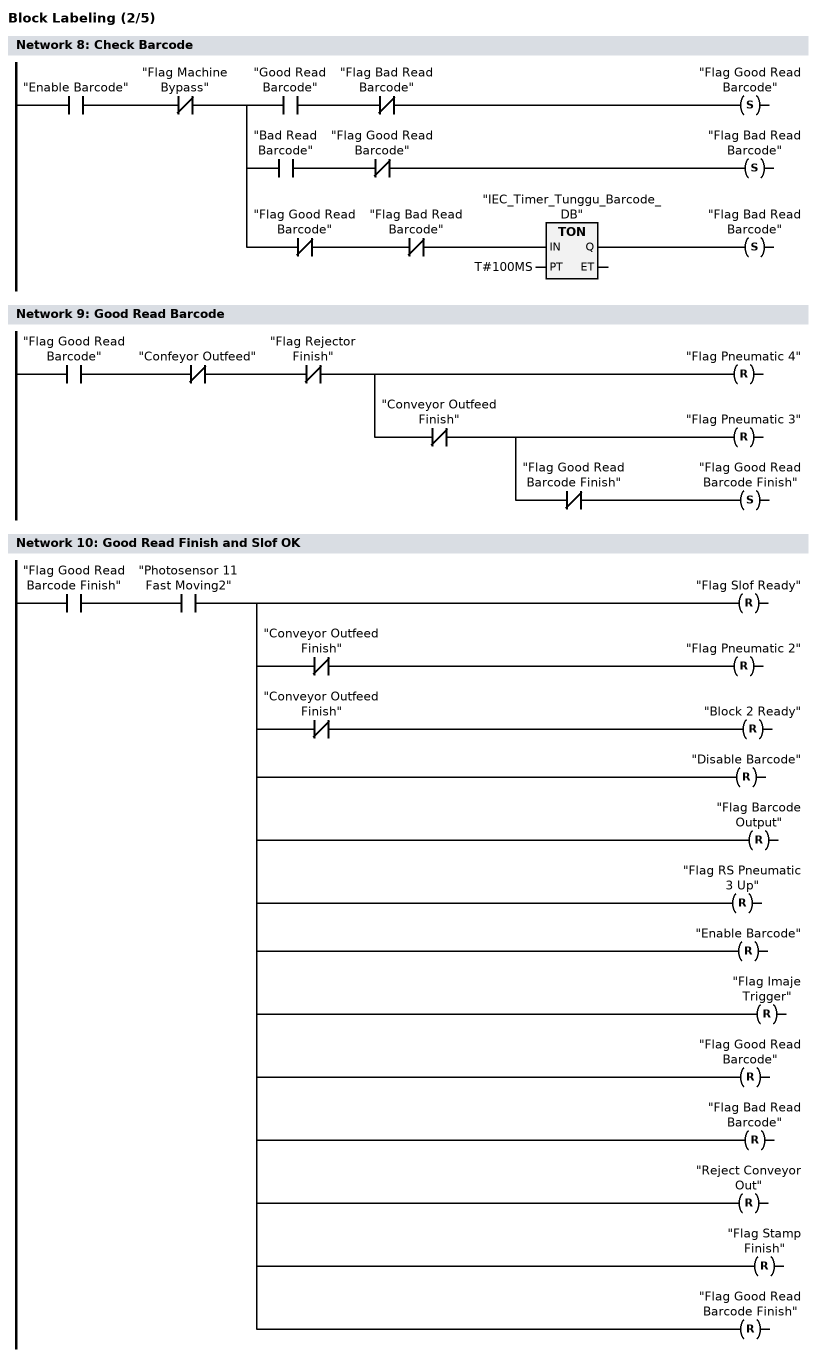
   #_w1 := "Enable Barcode" AND NOT "Flag Machine Bypass";
   IF #_w1 AND "Good Read Barcode" AND NOT "Flag Bad Read Barcode" THEN
       "Flag Good Read Barcode" := TRUE;
   END_IF;
   IF #_w1 AND "Bad Read Barcode" AND NOT "Flag Good Read Barcode" THEN
       "Flag Bad Read Barcode" := TRUE;
   END_IF;
   "IEC_Timer_Tunggu_Barcode_DB".TON(IN := #_w1 AND NOT "Flag Good Read Barcode" AND NOT "Flag Bad Read Barcode",
                           PT := T#100MS);
   IF "IEC_Timer_Tunggu_Barcode_DB".Q THEN "Flag Bad Read Barcode" := TRUE; END_IF;
END_REGION

REGION Network 9: Good Read Barcode
   RUNG wire#powerrail
      Contact( "Flag Good Read Barcode" )
      I_Contact( "Confeyor Outfeed" )
      I_Contact( "Flag Rejector Finish" )
      wire#w1
      R_Coil( "Flag Pneumatic 4" )
   END_RUNG
   RUNG wire#w1
      I_Contact( "Conveyor Outfeed Finish" )
      wire#w2
      R_Coil( "Flag Pneumatic 3" )
   END_RUNG
   RUNG wire#w2
      I_Contact( "Flag Good Read Barcode Finish" )
      S_Coil( "Flag Good Read Barcode Finish" )
   END_RUNG
   // the same network as SCL:
   #_w1 := "Flag Good Read Barcode" AND NOT "Confeyor Outfeed" AND NOT "Flag Rejector Finish";
   IF #_w1 THEN "Flag Pneumatic 4" := FALSE; END_IF;
   #_w2 := #_w1 AND NOT "Conveyor Outfeed Finish";
   IF #_w2 THEN "Flag Pneumatic 3" := FALSE; END_IF;
   IF #_w2 AND NOT "Flag Good Read Barcode Finish" THEN "Flag Good Read Barcode Finish" := TRUE; END_IF;
END_REGION

REGION Network 10: Good Read Finish and Slof OK
   RUNG wire#powerrail
      Contact( "Flag Good Read Barcode Finish" )
      Contact( "Photosensor 11 Fast Moving2" )
      wire#w1
      R_Coil( "Flag Slof Ready" )
   END_RUNG
   RUNG wire#w1
      I_Contact( "Conveyor Outfeed Finish" )
      R_Coil( "Flag Pneumatic 2" )
   END_RUNG
   RUNG wire#w1
      I_Contact( "Conveyor Outfeed Finish" )
      R_Coil( "Block 2 Ready" )
   END_RUNG
   RUNG wire#w1
      R_Coil( "Disable Barcode" )
   END_RUNG
   RUNG wire#w1
      R_Coil( "Flag Barcode Output" )
   END_RUNG
   RUNG wire#w1
      R_Coil( "Flag RS Pneumatic 3 Up" )
   END_RUNG
   RUNG wire#w1
      R_Coil( "Enable Barcode" )
   END_RUNG
   RUNG wire#w1
      R_Coil( "Flag Imaje Trigger" )
   END_RUNG
   RUNG wire#w1
      R_Coil( "Flag Good Read Barcode" )
   END_RUNG
   RUNG wire#w1
      R_Coil( "Flag Bad Read Barcode" )
   END_RUNG
   RUNG wire#w1
      R_Coil( "Reject Conveyor Out" )
   END_RUNG
   RUNG wire#w1
      R_Coil( "Flag Stamp Finish" )
   END_RUNG
   RUNG wire#w1
      R_Coil( "Flag Good Read Barcode Finish" )
   END_RUNG
   // the same network as SCL:
   #_w1 := "Flag Good Read Barcode Finish" AND "Photosensor 11 Fast Moving2";
   IF #_w1 THEN "Flag Slof Ready" := FALSE; END_IF;
   IF #_w1 AND NOT "Conveyor Outfeed Finish" THEN
       "Flag Pneumatic 2" := FALSE;
       "Block 2 Ready" := FALSE;
   END_IF;
   IF #_w1 THEN
       "Disable Barcode" := FALSE;
       "Flag Barcode Output" := FALSE;
       "Flag RS Pneumatic 3 Up" := FALSE;
       "Enable Barcode" := FALSE;
       "Flag Imaje Trigger" := FALSE;
       "Flag Good Read Barcode" := FALSE;
       "Flag Bad Read Barcode" := FALSE;
       "Reject Conveyor Out" := FALSE;
       "Flag Stamp Finish" := FALSE;
       "Flag Good Read Barcode Finish" := FALSE;
   END_IF;
END_REGION

REGION Network 11: Set Section Reject
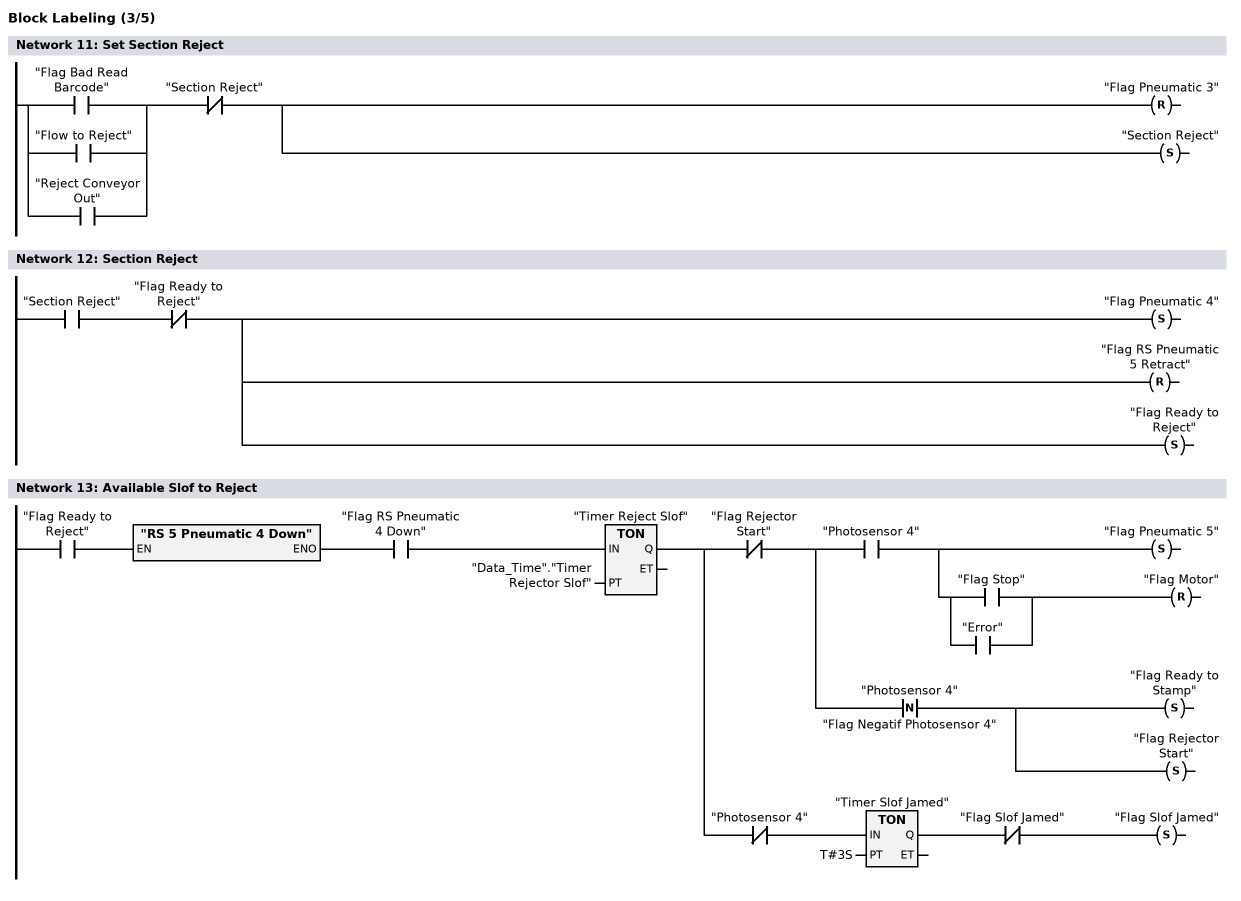
   RUNG wire#powerrail
      Contact( "Flag Bad Read Barcode" )
      wire#w1
      I_Contact( "Section Reject" )
      wire#w2
      R_Coil( "Flag Pneumatic 3" )
   END_RUNG
   RUNG wire#powerrail
      Contact( "Flow to Reject" )
   END_RUNG wire#w1
   RUNG wire#powerrail
      Contact( "Reject Conveyor Out" )
   END_RUNG wire#w1
   RUNG wire#w2
      S_Coil( "Section Reject" )
   END_RUNG
   // the same network as SCL:
   IF ("Flag Bad Read Barcode" OR "Flow to Reject" OR "Reject Conveyor Out") AND NOT "Section Reject" THEN
       "Flag Pneumatic 3" := FALSE;
       "Section Reject" := TRUE;
   END_IF;
END_REGION

REGION Network 12: Section Reject
   RUNG wire#powerrail
      Contact( "Section Reject" )
      I_Contact( "Flag Ready to Reject" )
      wire#w1
      S_Coil( "Flag Pneumatic 4" )
   END_RUNG
   RUNG wire#w1
      R_Coil( "Flag RS Pneumatic 5 Retract" )
   END_RUNG
   RUNG wire#w1
      S_Coil( "Flag Ready to Reject" )
   END_RUNG
   // the same network as SCL:
   IF "Section Reject" AND NOT "Flag Ready to Reject" THEN
       "Flag Pneumatic 4" := TRUE;
       "Flag RS Pneumatic 5 Retract" := FALSE;
       "Flag Ready to Reject" := TRUE;
   END_IF;
END_REGION

REGION Network 13: Available Slof to Reject
   "RS 5 Pneumatic 4 Down"(EN := "Flag Ready to Reject", ENO => #_w1);
   "Timer Reject Slof".TON(IN := #_w1 AND "Flag RS Pneumatic 4 Down", PT := "Data_Time"."Timer Rejector Slof");
   #_w2 := "Timer Reject Slof".Q AND NOT "Flag Rejector Start";
   #_w3 := #_w2 AND "Photosensor 4";
   IF #_w3 THEN "Flag Pneumatic 5" := TRUE; END_IF;
   IF #_w3 AND ("Flag Stop" OR "Error") THEN "Flag Motor" := FALSE; END_IF;
   #_w4 := #_w2 AND NOT "Photosensor 4" AND "Flag Negatif Photosensor 4";   // falling edge of "Photosensor 4"
   "Flag Negatif Photosensor 4" := "Photosensor 4";
   IF #_w4 THEN
       "Flag Ready to Stamp" := TRUE;
       "Flag Rejector Start" := TRUE;
   END_IF;
   "Timer Slof Jamed".TON(IN := "Timer Reject Slof".Q AND NOT "Photosensor 4", PT := T#3S);
   IF "Timer Slof Jamed".Q AND NOT "Flag Slof Jamed" THEN "Flag Slof Jamed" := TRUE; END_IF;
END_REGION

REGION Network 14: Ready to Stamp again
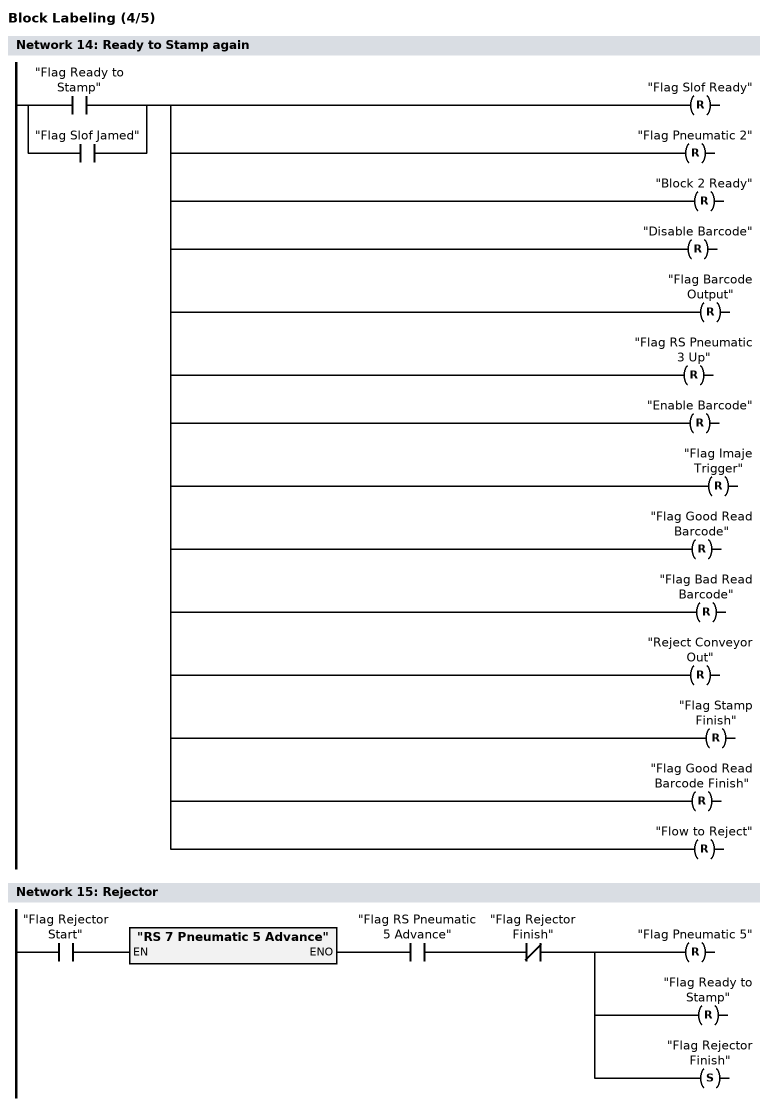
   RUNG wire#powerrail
      Contact( "Flag Ready to Stamp" )
      wire#w1
      R_Coil( "Flag Slof Ready" )
   END_RUNG
   RUNG wire#powerrail
      Contact( "Flag Slof Jamed" )
   END_RUNG wire#w1
   RUNG wire#w1
      R_Coil( "Flag Pneumatic 2" )
   END_RUNG
   RUNG wire#w1
      R_Coil( "Block 2 Ready" )
   END_RUNG
   RUNG wire#w1
      R_Coil( "Disable Barcode" )
   END_RUNG
   RUNG wire#w1
      R_Coil( "Flag Barcode Output" )
   END_RUNG
   RUNG wire#w1
      R_Coil( "Flag RS Pneumatic 3 Up" )
   END_RUNG
   RUNG wire#w1
      R_Coil( "Enable Barcode" )
   END_RUNG
   RUNG wire#w1
      R_Coil( "Flag Imaje Trigger" )
   END_RUNG
   RUNG wire#w1
      R_Coil( "Flag Good Read Barcode" )
   END_RUNG
   RUNG wire#w1
      R_Coil( "Flag Bad Read Barcode" )
   END_RUNG
   RUNG wire#w1
      R_Coil( "Reject Conveyor Out" )
   END_RUNG
   RUNG wire#w1
      R_Coil( "Flag Stamp Finish" )
   END_RUNG
   RUNG wire#w1
      R_Coil( "Flag Good Read Barcode Finish" )
   END_RUNG
   RUNG wire#w1
      R_Coil( "Flow to Reject" )
   END_RUNG
   // the same network as SCL:
   IF "Flag Ready to Stamp" OR "Flag Slof Jamed" THEN
       "Flag Slof Ready" := FALSE;
       "Flag Pneumatic 2" := FALSE;
       "Block 2 Ready" := FALSE;
       "Disable Barcode" := FALSE;
       "Flag Barcode Output" := FALSE;
       "Flag RS Pneumatic 3 Up" := FALSE;
       "Enable Barcode" := FALSE;
       "Flag Imaje Trigger" := FALSE;
       "Flag Good Read Barcode" := FALSE;
       "Flag Bad Read Barcode" := FALSE;
       "Reject Conveyor Out" := FALSE;
       "Flag Stamp Finish" := FALSE;
       "Flag Good Read Barcode Finish" := FALSE;
       "Flow to Reject" := FALSE;
   END_IF;
END_REGION

REGION Network 15: Rejector
   RUNG wire#powerrail
      Contact( "Flag Rejector Start" )
      "RS 7 Pneumatic 5 Advance"()
      Contact( "Flag RS Pneumatic 5 Advance" )
      I_Contact( "Flag Rejector Finish" )
      wire#w1
      R_Coil( "Flag Pneumatic 5" )
   END_RUNG
   RUNG wire#w1
      R_Coil( "Flag Ready to Stamp" )
   END_RUNG
   RUNG wire#w1
      S_Coil( "Flag Rejector Finish" )
   END_RUNG
   // the same network as SCL:
   "RS 7 Pneumatic 5 Advance"(EN := "Flag Rejector Start", ENO => #_w1);
   IF #_w1 AND "Flag RS Pneumatic 5 Advance" AND NOT "Flag Rejector Finish" THEN
       "Flag Pneumatic 5" := FALSE;
       "Flag Ready to Stamp" := FALSE;
       "Flag Rejector Finish" := TRUE;
   END_IF;
END_REGION

REGION Network 16: Rejector Finish
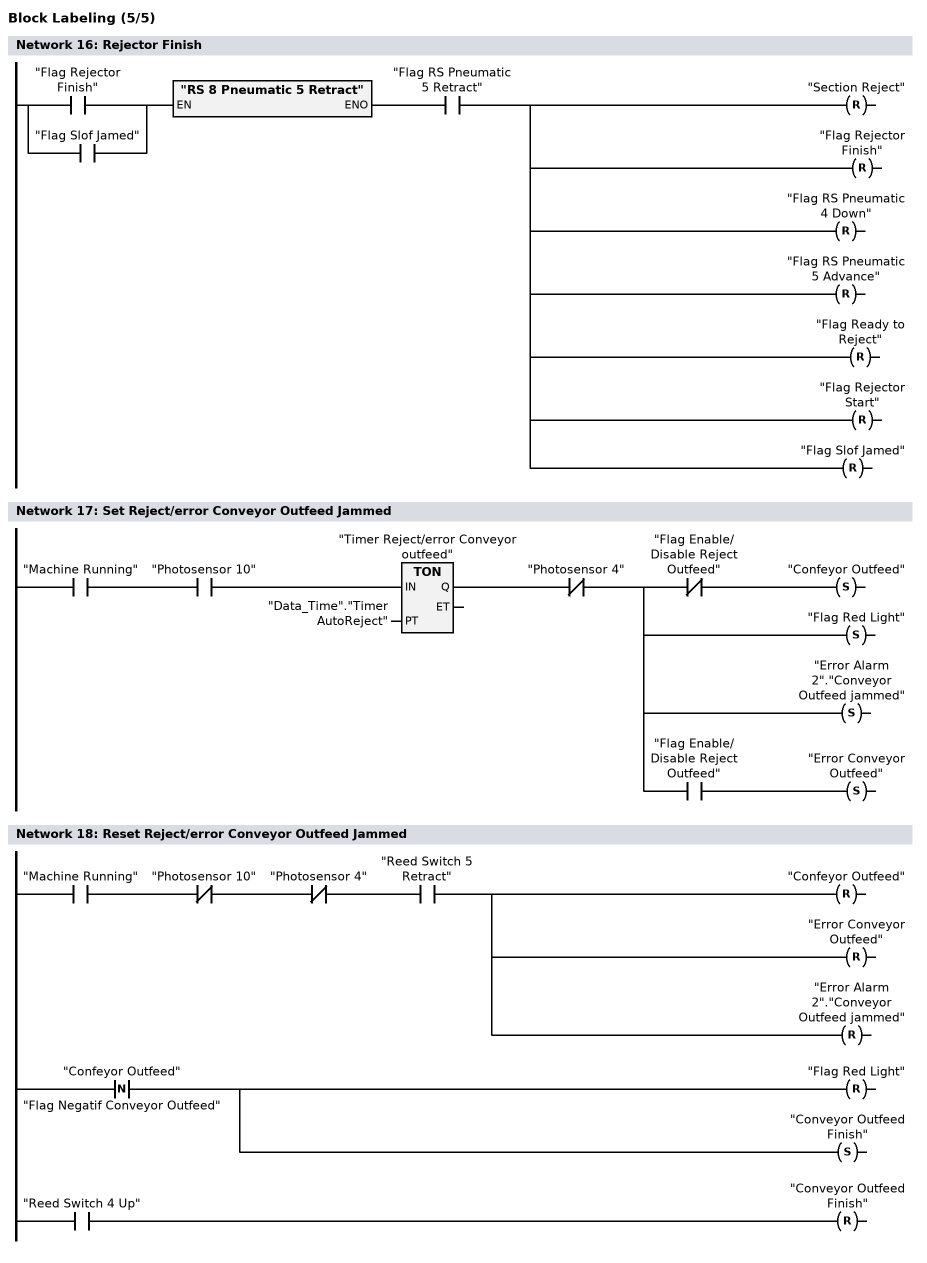
   RUNG wire#powerrail
      Contact( "Flag Rejector Finish" )
      wire#w1
      "RS 8 Pneumatic 5 Retract"()
      Contact( "Flag RS Pneumatic 5 Retract" )
      wire#w2
      R_Coil( "Section Reject" )
   END_RUNG
   RUNG wire#powerrail
      Contact( "Flag Slof Jamed" )
   END_RUNG wire#w1
   RUNG wire#w2
      R_Coil( "Flag Rejector Finish" )
   END_RUNG
   RUNG wire#w2
      R_Coil( "Flag RS Pneumatic 4 Down" )
   END_RUNG
   RUNG wire#w2
      R_Coil( "Flag RS Pneumatic 5 Advance" )
   END_RUNG
   RUNG wire#w2
      R_Coil( "Flag Ready to Reject" )
   END_RUNG
   RUNG wire#w2
      R_Coil( "Flag Rejector Start" )
   END_RUNG
   RUNG wire#w2
      R_Coil( "Flag Slof Jamed" )
   END_RUNG
   // the same network as SCL:
   "RS 8 Pneumatic 5 Retract"(EN := "Flag Rejector Finish" OR "Flag Slof Jamed", ENO => #_w1);
   IF #_w1 AND "Flag RS Pneumatic 5 Retract" THEN
       "Section Reject" := FALSE;
       "Flag Rejector Finish" := FALSE;
       "Flag RS Pneumatic 4 Down" := FALSE;
       "Flag RS Pneumatic 5 Advance" := FALSE;
       "Flag Ready to Reject" := FALSE;
       "Flag Rejector Start" := FALSE;
       "Flag Slof Jamed" := FALSE;
   END_IF;
END_REGION

REGION Network 17: Set Reject/error Conveyor Outfeed Jammed
   "Timer Reject/error Conveyor outfeed".TON(IN := "Machine Running" AND "Photosensor 10",
                           PT := "Data_Time"."Timer AutoReject");
   #_w1 := "Timer Reject/error Conveyor outfeed".Q AND NOT "Photosensor 4";
   IF #_w1 AND NOT "Flag Enable/Disable Reject Outfeed" THEN "Confeyor Outfeed" := TRUE; END_IF;
   IF #_w1 THEN
       "Flag Red Light" := TRUE;
       "Error Alarm 2"."Conveyor Outfeed jammed" := TRUE;
   END_IF;
   IF #_w1 AND "Flag Enable/Disable Reject Outfeed" THEN "Error Conveyor Outfeed" := TRUE; END_IF;
END_REGION

REGION Network 18: Reset Reject/error Conveyor Outfeed Jammed
   RUNG wire#powerrail
      Contact( "Machine Running" )
      I_Contact( "Photosensor 10" )
      I_Contact( "Photosensor 4" )
      Contact( "Reed Switch 5 Retract" )
      wire#w1
      R_Coil( "Confeyor Outfeed" )
   END_RUNG
   RUNG wire#w1
      R_Coil( "Error Conveyor Outfeed" )
   END_RUNG
   RUNG wire#w1
      R_Coil( "Error Alarm 2"."Conveyor Outfeed jammed" )
   END_RUNG
   RUNG wire#powerrail
      N_Contact(operand := "Confeyor Outfeed", bit := "Flag Negatif Conveyor Outfeed")
      wire#w2
      R_Coil( "Flag Red Light" )
   END_RUNG
   RUNG wire#w2
      S_Coil( "Conveyor Outfeed Finish" )
   END_RUNG
   RUNG wire#powerrail
      Contact( "Reed Switch 4 Up" )
      R_Coil( "Conveyor Outfeed Finish" )
   END_RUNG
   // the same network as SCL:
   IF "Machine Running" AND NOT "Photosensor 10" AND NOT "Photosensor 4" AND "Reed Switch 5 Retract" THEN
       "Confeyor Outfeed" := FALSE;
       "Error Conveyor Outfeed" := FALSE;
       "Error Alarm 2"."Conveyor Outfeed jammed" := FALSE;
   END_IF;
   #_w1 := NOT "Confeyor Outfeed" AND "Flag Negatif Conveyor Outfeed";   // falling edge of "Confeyor Outfeed"
   "Flag Negatif Conveyor Outfeed" := "Confeyor Outfeed";
   IF #_w1 THEN
       "Flag Red Light" := FALSE;
       "Conveyor Outfeed Finish" := TRUE;
   END_IF;
   IF "Reed Switch 4 Up" THEN "Conveyor Outfeed Finish" := FALSE; END_IF;
END_REGION
END_FUNCTION_BLOCK

FUNCTION_BLOCK "Block Focke"   // FB6, LAD
{ S7_Optimized_Access := 'TRUE' }
VERSION : 0.1
   VAR_TEMP   // added for the SCL form of the ladder/FBD networks
      _w1 : Bool;
   END_VAR
BEGIN

REGION Network 1: Enable/Disable Error Chute Before Heating Roll
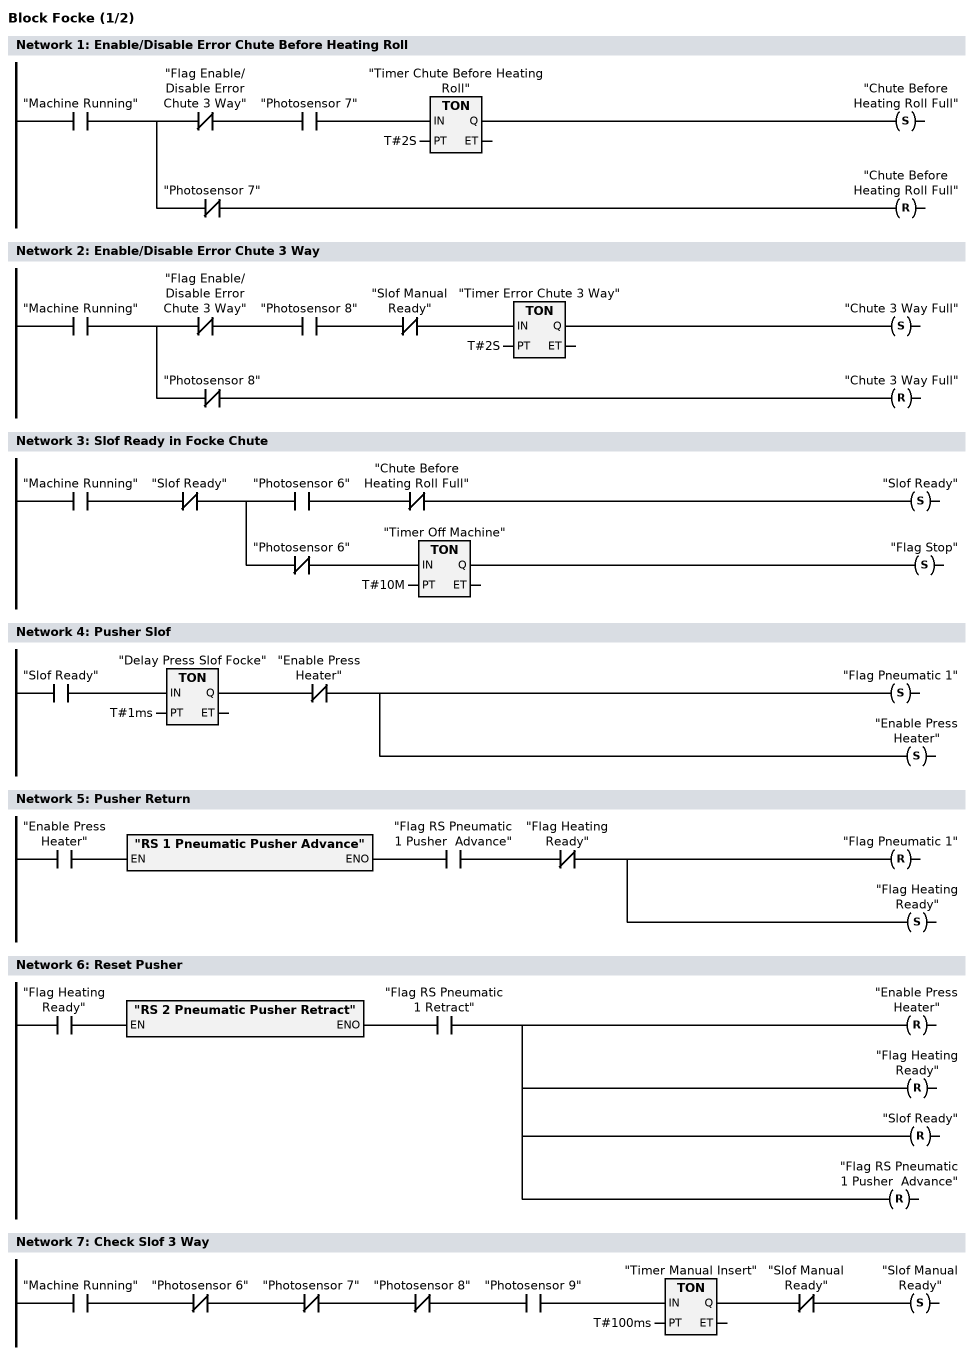
   "Timer Chute Before Heating Roll".TON(IN := "Machine Running" AND NOT "Flag Enable/Disable Error Chute 3 Way" AND "Photosensor 7",
                           PT := T#2S);
   IF "Timer Chute Before Heating Roll".Q THEN "Chute Before Heating Roll Full" := TRUE; END_IF;
   IF "Machine Running" AND NOT "Photosensor 7" THEN "Chute Before Heating Roll Full" := FALSE; END_IF;
END_REGION

REGION Network 2: Enable/Disable Error Chute 3 Way
   "Timer Error Chute 3 Way".TON(IN := "Machine Running" AND NOT "Flag Enable/Disable Error Chute 3 Way" AND "Photosensor 8" AND NOT "Slof Manual Ready",
                           PT := T#2S);
   IF "Timer Error Chute 3 Way".Q THEN "Chute 3 Way Full" := TRUE; END_IF;
   IF "Machine Running" AND NOT "Photosensor 8" THEN "Chute 3 Way Full" := FALSE; END_IF;
END_REGION

REGION Network 3: Slof Ready in Focke Chute
   #_w1 := "Machine Running" AND NOT "Slof Ready";
   IF #_w1 AND "Photosensor 6" AND NOT "Chute Before Heating Roll Full" THEN "Slof Ready" := TRUE; END_IF;
   "Timer Off Machine".TON(IN := #_w1 AND NOT "Photosensor 6", PT := T#10M);
   IF "Timer Off Machine".Q THEN "Flag Stop" := TRUE; END_IF;
END_REGION

REGION Network 4: Pusher Slof
   "Delay Press Slof Focke".TON(IN := "Slof Ready", PT := T#1ms);
   IF "Delay Press Slof Focke".Q AND NOT "Enable Press Heater" THEN
       "Flag Pneumatic 1" := TRUE;
       "Enable Press Heater" := TRUE;
   END_IF;
END_REGION

REGION Network 5: Pusher Return
   RUNG wire#powerrail
      Contact( "Enable Press Heater" )
      "RS 1 Pneumatic Pusher Advance"()
      Contact( "Flag RS Pneumatic 1 Pusher  Advance" )
      I_Contact( "Flag Heating Ready" )
      wire#w1
      R_Coil( "Flag Pneumatic 1" )
   END_RUNG
   RUNG wire#w1
      S_Coil( "Flag Heating Ready" )
   END_RUNG
   // the same network as SCL:
   "RS 1 Pneumatic Pusher Advance"(EN := "Enable Press Heater", ENO => #_w1);
   IF #_w1 AND "Flag RS Pneumatic 1 Pusher  Advance" AND NOT "Flag Heating Ready" THEN
       "Flag Pneumatic 1" := FALSE;
       "Flag Heating Ready" := TRUE;
   END_IF;
END_REGION

REGION Network 6: Reset Pusher
   RUNG wire#powerrail
      Contact( "Flag Heating Ready" )
      "RS 2 Pneumatic Pusher Retract"()
      Contact( "Flag RS Pneumatic 1 Retract" )
      wire#w1
      R_Coil( "Enable Press Heater" )
   END_RUNG
   RUNG wire#w1
      R_Coil( "Flag Heating Ready" )
   END_RUNG
   RUNG wire#w1
      R_Coil( "Slof Ready" )
   END_RUNG
   RUNG wire#w1
      R_Coil( "Flag RS Pneumatic 1 Pusher  Advance" )
   END_RUNG
   // the same network as SCL:
   "RS 2 Pneumatic Pusher Retract"(EN := "Flag Heating Ready", ENO => #_w1);
   IF #_w1 AND "Flag RS Pneumatic 1 Retract" THEN
       "Enable Press Heater" := FALSE;
       "Flag Heating Ready" := FALSE;
       "Slof Ready" := FALSE;
       "Flag RS Pneumatic 1 Pusher  Advance" := FALSE;
   END_IF;
END_REGION

REGION Network 7: Check Slof 3 Way
   "Timer Manual Insert".TON(IN := "Machine Running" AND NOT "Photosensor 6" AND NOT "Photosensor 7" AND NOT "Photosensor 8" AND "Photosensor 9",
                           PT := T#100ms);
   IF "Timer Manual Insert".Q AND NOT "Slof Manual Ready" THEN "Slof Manual Ready" := TRUE; END_IF;
END_REGION

REGION Network 8: Manual Insert Slof
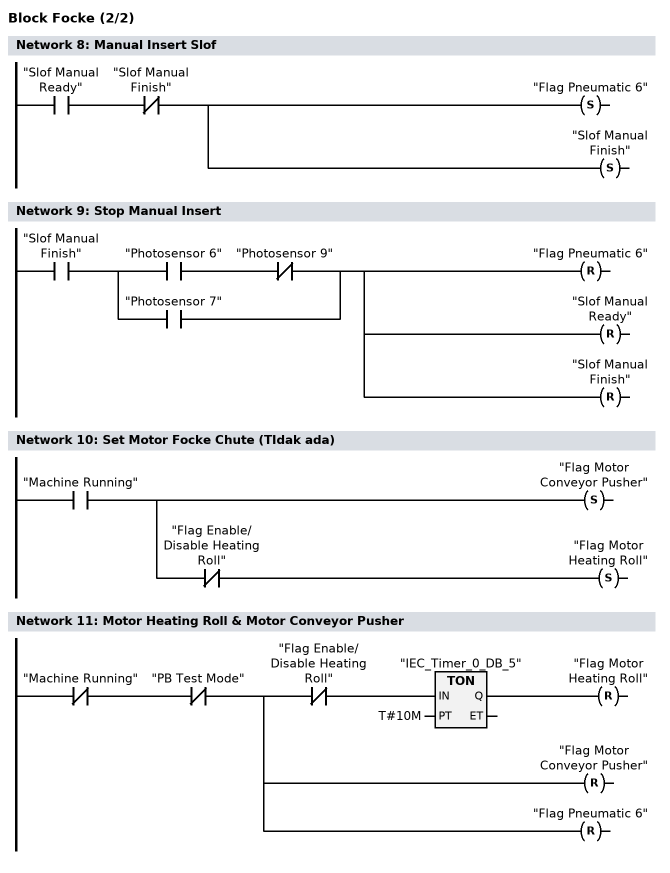
   RUNG wire#powerrail
      Contact( "Slof Manual Ready" )
      I_Contact( "Slof Manual Finish" )
      wire#w1
      S_Coil( "Flag Pneumatic 6" )
   END_RUNG
   RUNG wire#w1
      S_Coil( "Slof Manual Finish" )
   END_RUNG
   // the same network as SCL:
   IF "Slof Manual Ready" AND NOT "Slof Manual Finish" THEN
       "Flag Pneumatic 6" := TRUE;
       "Slof Manual Finish" := TRUE;
   END_IF;
END_REGION

REGION Network 9: Stop Manual Insert
   RUNG wire#powerrail
      Contact( "Slof Manual Finish" )
      wire#w1
      Contact( "Photosensor 6" )
      I_Contact( "Photosensor 9" )
      wire#w2
      R_Coil( "Flag Pneumatic 6" )
   END_RUNG
   RUNG wire#w1
      Contact( "Photosensor 7" )
   END_RUNG wire#w2
   RUNG wire#w2
      R_Coil( "Slof Manual Ready" )
   END_RUNG
   RUNG wire#w2
      R_Coil( "Slof Manual Finish" )
   END_RUNG
   // the same network as SCL:
   IF "Slof Manual Finish" AND (("Photosensor 6" AND NOT "Photosensor 9") OR "Photosensor 7") THEN
       "Flag Pneumatic 6" := FALSE;
       "Slof Manual Ready" := FALSE;
       "Slof Manual Finish" := FALSE;
   END_IF;
END_REGION

REGION Network 10: Set Motor Focke Chute (TIdak ada)
   RUNG wire#powerrail
      Contact( "Machine Running" )
      wire#w1
      S_Coil( "Flag Motor Conveyor Pusher" )
   END_RUNG
   RUNG wire#w1
      I_Contact( "Flag Enable/Disable Heating Roll" )
      S_Coil( "Flag Motor Heating Roll" )
   END_RUNG
   // the same network as SCL:
   IF "Machine Running" THEN "Flag Motor Conveyor Pusher" := TRUE; END_IF;
   IF "Machine Running" AND NOT "Flag Enable/Disable Heating Roll" THEN
       "Flag Motor Heating Roll" := TRUE;
   END_IF;
END_REGION

REGION Network 11: Motor Heating Roll & Motor Conveyor Pusher
   #_w1 := NOT "Machine Running" AND NOT "PB Test Mode";
   "IEC_Timer_0_DB_5".TON(IN := #_w1 AND NOT "Flag Enable/Disable Heating Roll", PT := T#10M);
   IF "IEC_Timer_0_DB_5".Q THEN "Flag Motor Heating Roll" := FALSE; END_IF;
   IF #_w1 THEN
       "Flag Motor Conveyor Pusher" := FALSE;
       "Flag Pneumatic 6" := FALSE;
   END_IF;
END_REGION
END_FUNCTION_BLOCK

FUNCTION_BLOCK "S Block Par Statistika"   // FB7, LAD
{ S7_Optimized_Access := 'TRUE' }
VERSION : 0.1
BEGIN

REGION Network 1: Move Data Dari HMI Ke Setting Time
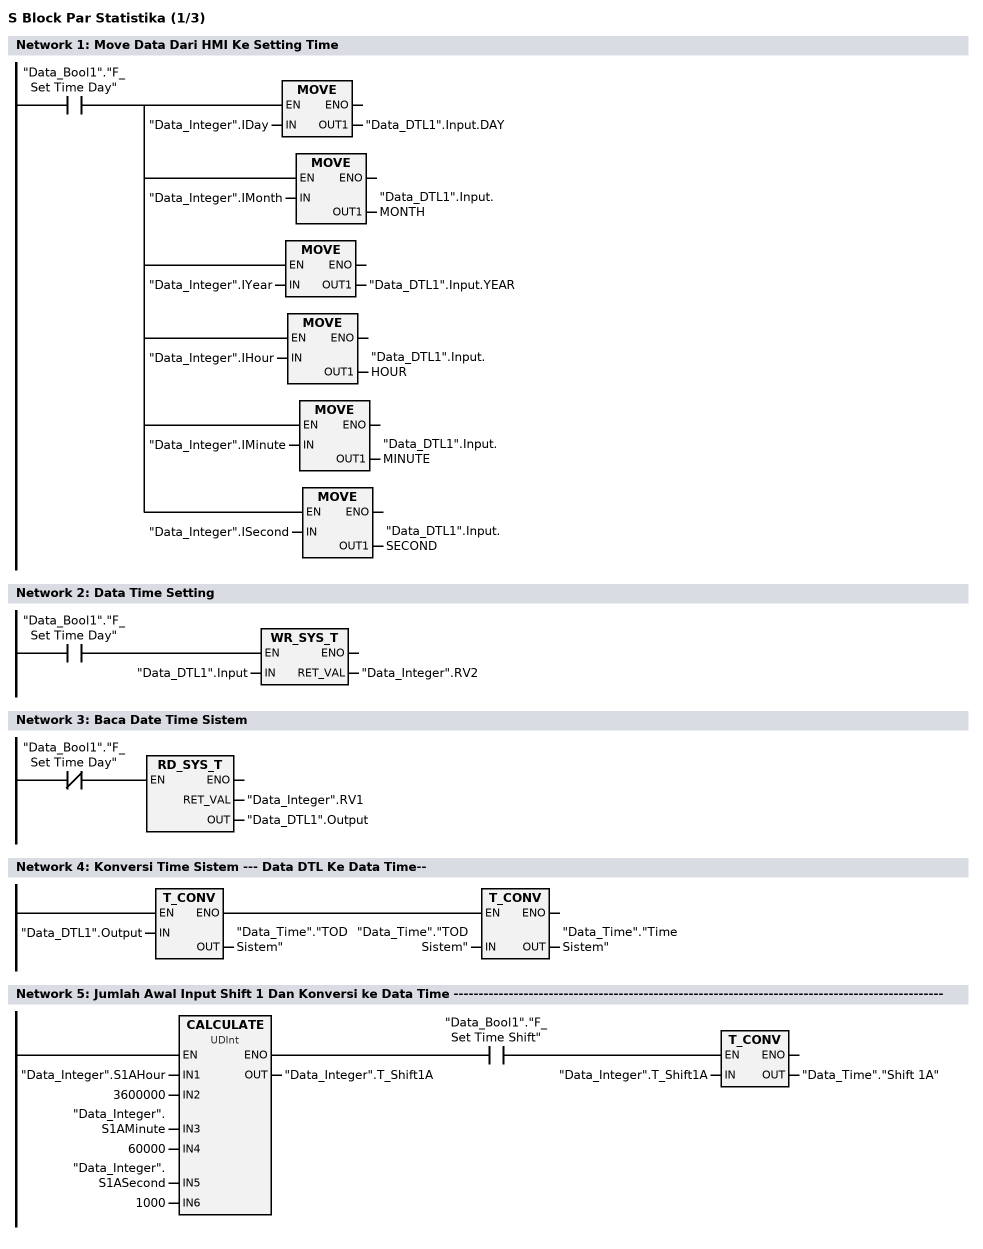
   RUNG wire#powerrail
      Contact( "Data_Bool1"."F_Set Time Day" )
      wire#w1
      { S7_GenerateENO := "TRUE" } Move(in := "Data_Integer".IDay, out1 => "Data_DTL1".Input.DAY)
   END_RUNG
   RUNG wire#w1
      { S7_GenerateENO := "TRUE" } Move(in := "Data_Integer".IMonth, out1 => "Data_DTL1".Input.MONTH)
   END_RUNG
   RUNG wire#w1
      { S7_GenerateENO := "TRUE" } Move(in := "Data_Integer".IYear, out1 => "Data_DTL1".Input.YEAR)
   END_RUNG
   RUNG wire#w1
      { S7_GenerateENO := "TRUE" } Move(in := "Data_Integer".IHour, out1 => "Data_DTL1".Input.HOUR)
   END_RUNG
   RUNG wire#w1
      { S7_GenerateENO := "TRUE" } Move(in := "Data_Integer".IMinute, out1 => "Data_DTL1".Input.MINUTE)
   END_RUNG
   RUNG wire#w1
      { S7_GenerateENO := "TRUE" } Move(in := "Data_Integer".ISecond, out1 => "Data_DTL1".Input.SECOND)
   END_RUNG
   // the same network as SCL:
   IF "Data_Bool1"."F_Set Time Day" THEN
       "Data_DTL1".Input.DAY := "Data_Integer".IDay;
       "Data_DTL1".Input.MONTH := "Data_Integer".IMonth;
       "Data_DTL1".Input.YEAR := "Data_Integer".IYear;
       "Data_DTL1".Input.HOUR := "Data_Integer".IHour;
       "Data_DTL1".Input.MINUTE := "Data_Integer".IMinute;
       "Data_DTL1".Input.SECOND := "Data_Integer".ISecond;
   END_IF;
END_REGION

REGION Network 2: Data Time Setting
   IF "Data_Bool1"."F_Set Time Day" THEN "Data_Integer".RV2 := WR_SYS_T(IN := "Data_DTL1".Input); END_IF;
END_REGION

REGION Network 3: Baca Date Time Sistem
   IF NOT "Data_Bool1"."F_Set Time Day" THEN
       "Data_Integer".RV1 := RD_SYS_T(OUT => "Data_DTL1".Output);
   END_IF;
END_REGION

REGION Network 4: Konversi Time Sistem --- Data DTL Ke Data Time--
   // ENO of a box is taken as its EN; it also drops when the box reports an error
   "Data_Time"."TOD Sistem" := T_CONV(IN := "Data_DTL1".Output);
   "Data_Time"."Time Sistem" := T_CONV(IN := "Data_Time"."TOD Sistem");
END_REGION

REGION Network 5: Jumlah Awal Input Shift 1 Dan Konversi ke Data Time --------------------------------------------------------------------------------------------------
   // ENO of a box is taken as its EN; it also drops when the box reports an error
   "Data_Integer".T_Shift1A := ("Data_Integer".S1AHour*3600000)+("Data_Integer".S1AMinute*60000)+("Data_Integer".S1ASecond*1000);
   IF "Data_Bool1"."F_Set Time Shift" THEN
       "Data_Time"."Shift 1A" := T_CONV(IN := "Data_Integer".T_Shift1A);
   END_IF;
END_REGION

REGION Network 6: Jumlah Akhir Input Shift 1 Dan Konversi ke Data Time @@@@@@@@@@@
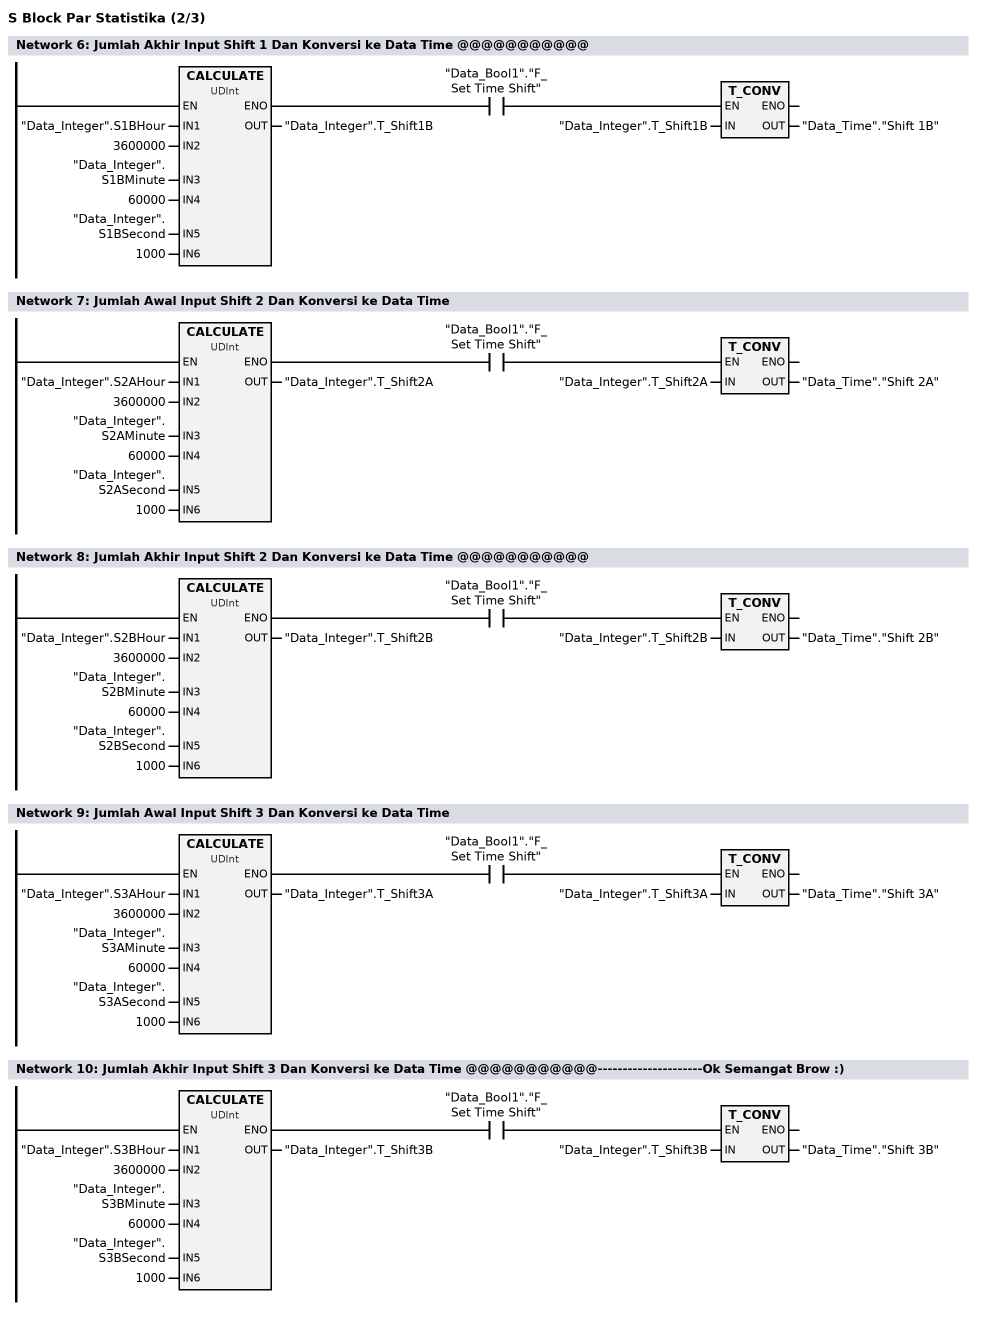
   // ENO of a box is taken as its EN; it also drops when the box reports an error
   "Data_Integer".T_Shift1B := ("Data_Integer".S1BHour*3600000)+("Data_Integer".S1BMinute*60000)+("Data_Integer".S1BSecond*1000);
   IF "Data_Bool1"."F_Set Time Shift" THEN
       "Data_Time"."Shift 1B" := T_CONV(IN := "Data_Integer".T_Shift1B);
   END_IF;
END_REGION

REGION Network 7: Jumlah Awal Input Shift 2 Dan Konversi ke Data Time
   // ENO of a box is taken as its EN; it also drops when the box reports an error
   "Data_Integer".T_Shift2A := ("Data_Integer".S2AHour*3600000)+("Data_Integer".S2AMinute*60000)+("Data_Integer".S2ASecond*1000);
   IF "Data_Bool1"."F_Set Time Shift" THEN
       "Data_Time"."Shift 2A" := T_CONV(IN := "Data_Integer".T_Shift2A);
   END_IF;
END_REGION

REGION Network 8: Jumlah Akhir Input Shift 2 Dan Konversi ke Data Time @@@@@@@@@@@
   // ENO of a box is taken as its EN; it also drops when the box reports an error
   "Data_Integer".T_Shift2B := ("Data_Integer".S2BHour*3600000)+("Data_Integer".S2BMinute*60000)+("Data_Integer".S2BSecond*1000);
   IF "Data_Bool1"."F_Set Time Shift" THEN
       "Data_Time"."Shift 2B" := T_CONV(IN := "Data_Integer".T_Shift2B);
   END_IF;
END_REGION

REGION Network 9: Jumlah Awal Input Shift 3 Dan Konversi ke Data Time
   // ENO of a box is taken as its EN; it also drops when the box reports an error
   "Data_Integer".T_Shift3A := ("Data_Integer".S3AHour*3600000)+("Data_Integer".S3AMinute*60000)+("Data_Integer".S3ASecond*1000);
   IF "Data_Bool1"."F_Set Time Shift" THEN
       "Data_Time"."Shift 3A" := T_CONV(IN := "Data_Integer".T_Shift3A);
   END_IF;
END_REGION

REGION Network 10: Jumlah Akhir Input Shift 3 Dan Konversi ke Data Time @@@@@@@@@@@---------------------Ok Semangat Brow :)
   // ENO of a box is taken as its EN; it also drops when the box reports an error
   "Data_Integer".T_Shift3B := ("Data_Integer".S3BHour*3600000)+("Data_Integer".S3BMinute*60000)+("Data_Integer".S3BSecond*1000);
   IF "Data_Bool1"."F_Set Time Shift" THEN
       "Data_Time"."Shift 3B" := T_CONV(IN := "Data_Integer".T_Shift3B);
   END_IF;
END_REGION

REGION Network 11: Data Time 5 Detik Sebelum Akhir Shift (Waktu Proses Copy Data Current minus 1 sampai 5
